(* Logix 5000 project; controller PLC_MCC1300_75F1 vendor 1 type 14 code 166 rev 32.11; software revision 32.04; part 81 of 83 *)
(* tags used below, declared in another part *)
   GP_OB_InitializeMain : GP_OB_Initialize;
   M302SpeedUp : MAC_SpeedUp;
   M307D_M1_DR : AXIS_CIP_DRIVE;
   M307E_M1_DR : AXIS_CIP_DRIVE;
   M307F_M1_DR : AXIS_CIP_DRIVE;
   M310_M1_DR_R1 : AXIS_CIP_DRIVE;
   M310_M2_DR_R2 : AXIS_CIP_DRIVE;
   M310_M3_DR_R3 : AXIS_CIP_DRIVE;
   TMP_dDirection : DINT;
   TMP_dTarget : DINT;
   TMP_rAcc : REAL;
   TMP_rDec : REAL;
   TMP_rSpeed : REAL;
   Z300_Conveyor : UDT_StandConv[29];
   Z300_Conveyor_IN_MOTION : MAC_Conveyor_ZC_IN_MOTION[29];
   Z300_Conveyor_OUT_MOTION : MAC_Conveyor_ZC_OUT_MOTION[29];
(* MotionLogic, continued *)

ROUTINE M307D_Motion   (* ladder *)
   // M307DM1
   0: NOP();
   1: XIC(Z300_Conveyor[18].OUTPUT_xDriveReset.0)MASR(M307D_M1_DR,Z300_Conveyor_OUT_MOTION[18].DR_MASR_M[0]);
   2: [XIC(Z300_Conveyor[18].OUTPUT_xDriveEnable.[0]) XIO(Z300_Conveyor_OUT_MOTION[18].DR_MSO_M[0].ER) MSO(M307D_M1_DR,Z300_Conveyor_OUT_MOTION[18].DR_MSO_M[0]) ,XIO(Z300_Conveyor_OUT_MOTION[18].DR_MSO_M[0].EN) OTU(Z300_Conveyor_OUT_MOTION[18].DR_MSO_M[0].ER) ,XIO(Z300_Conveyor[18].OUTPUT_xDriveEnable.[0]) OTU(Z300_Conveyor_OUT_MOTION[18].DR_MSO_M[0].EN) XIO(Z300_Conveyor_OUT_MOTION[18].DR_MSF_M[0].ER) MSF(M307D_M1_DR,Z300_Conveyor_OUT_MOTION[18].DR_MSF_M[0]) ,XIO(Z300_Conveyor_OUT_MOTION[18].DR_MSF_M[0].EN) OTU(Z300_Conveyor_OUT_MOTION[18].DR_MSF_M[0].ER) ];
   3: MUL(Z300_Conveyor[18].AUX_rgrAcc_m_s2[0],1000,TMP_rAcc)MUL(Z300_Conveyor[18].AUX_rgrDec_m_s2[0],1000,TMP_rDec)DIV(Z300_Conveyor[18].AUX_rgdRequestSpeed_mm_min[0],60,TMP_rSpeed);
   4: XIC(Z300_Conveyor[18].OS_xStartCount.0)OTU(Z300_Conveyor_IN_MOTION[18].DR_MAR_M[0].PC)OTU(Z300_Conveyor_IN_MOTION[18].DR_MRP_M[0].DN);
   5: [XIC(Z300_Conveyor[18].OUTPUT_xRun.0) MOV(0,TMP_dDirection) ,XIC(Z300_Conveyor[18].OUTPUT_xReverse.0) MOV(1,TMP_dDirection) ][XIO(Z300_Conveyor_IN_MOTION[18].DR_MAR_M[0].PC) ,XIO(Z300_Conveyor_IN_MOTION[18].DR_MRP_M[0].DN) ,XIO(Z300_Conveyor[18].OUTPUT_xPositioning.0) ]MAJ(M307D_M1_DR,Z300_Conveyor_OUT_MOTION[18].DR_MAJ_M[0],TMP_dDirection,TMP_rSpeed,Units per sec,TMP_rAcc,Units per sec2,TMP_rDec,Units per sec2,Trapezoidal,TMP_rAcc,TMP_rDec,Units per sec3,Enabled,Programmed,0,None);
   6: XIC(Z300_Conveyor[18].OS_xStartCount.0)MRP(M307D_M1_DR,Z300_Conveyor_OUT_MOTION[18].DR_MRP_M[0],Absolute,Actual,0);
   7: [XIC(Z300_Conveyor_IN_MOTION[18].DR_MRP_M[0].DN) XIC(Z300_Conveyor[18].OUTPUT_xPositioning.0) [XIC(Z300_Conveyor[18].tmON_PhFilter[0].DN) ,XIC(Z300_Conveyor_IN_MOTION[18].DR_MAR_M[0].EN) ] MAR(M307D_M1_DR,Z300_Conveyor_OUT_MOTION[18].DR_MAR_M[0],Negative_Edge,Disabled,0,0,1) ,XIO(Z300_Conveyor[18].OUTPUT_xPositioning.0) MDR(M307D_M1_DR,Z300_Conveyor_OUT_MOTION[18].DR_MDR_M[0],1) ];
   8: XIC(Z300_Conveyor[18].OUTPUT_xPositioning.0)XIC(Z300_Conveyor_IN_MOTION[18].DR_MAR_M[0].PC)DIV(Z300_Conveyor[18].AUX_rgdTarget_cmm[0],100,TMP_dTarget)ADD(TMP_dTarget,M307D_M1_DR.Registration1Position,TMP_dTarget)MAM(M307D_M1_DR,Z300_Conveyor_OUT_MOTION[18].DR_MAM_M[0],0,TMP_dTarget,TMP_rSpeed,Units per sec,TMP_rAcc,Units per sec2,TMP_rDec,Units per sec2,Trapezoidal,TMP_rAcc,TMP_rDec,Units per sec3,Enabled,Programmed,0,None,0,0);
   9: [XIC(Z300_Conveyor[18].OUTPUT_xChangeSpeed.0) ,XIC(M302SpeedUp.OS_xChangeAccDec) ,XIC(GP_OB_InitializeMain.OUT_xOs_200ms) ][XIO(Z300_Conveyor[18].OUTPUT_xReverse.0) ,XIC(Z300_Conveyor[18].OUTPUT_xReverse.0) MUL(TMP_rSpeed,-1.0,TMP_rSpeed) ]MCD(M307D_M1_DR,Z300_Conveyor_OUT_MOTION[18].DR_MCD_M[0],Jog,Yes,TMP_rSpeed,Yes,TMP_rAcc,Yes,TMP_rDec,No,TMP_rAcc,No,TMP_rDec,Units per sec,Units per sec2,Units per sec2,Units per sec3);
   10: XIO(Z300_Conveyor[18].OUTPUT_xRun.0)XIO(Z300_Conveyor[18].OUTPUT_xReverse.0)[XIC(Z300_Conveyor_IN_MOTION[18].DR_MAJ_M[0].IP) MAS(M307D_M1_DR,Z300_Conveyor_OUT_MOTION[18].DR_MASjog_M[0],Jog,Yes,TMP_rDec,Units per sec2,No,TMP_rDec,Units per sec3) ,XIC(Z300_Conveyor_IN_MOTION[18].DR_MAM_M[0].IP) MAS(M307D_M1_DR,Z300_Conveyor_OUT_MOTION[18].DR_MASpos_M[0],Move,Yes,TMP_rDec,Units per sec2,No,TMP_rDec,Units per sec3) ,XIO(Z300_Conveyor_IN_MOTION[18].DR_MAJ_M[0].IP) XIO(Z300_Conveyor_IN_MOTION[18].DR_MAM_M[0].IP) XIO(Z300_Conveyor_IN_MOTION[18].DR_MASjog_M[0].IP) XIO(Z300_Conveyor_IN_MOTION[18].DR_MASpos_M[0].IP) MAS(M307D_M1_DR,Z300_Conveyor_OUT_MOTION[18].DR_MASall_M[0],All,Yes,TMP_rDec,Units per sec2,No,TMP_rDec,Units per sec3) ];
END_ROUTINE

ROUTINE M307E_Motion   (* ladder *)
   // M307EM1
   0: NOP();
   1: XIC(Z300_Conveyor[19].OUTPUT_xDriveReset.0)MASR(M307E_M1_DR,Z300_Conveyor_OUT_MOTION[19].DR_MASR_M[0]);
   2: [XIC(Z300_Conveyor[19].OUTPUT_xDriveEnable.[0]) XIO(Z300_Conveyor_OUT_MOTION[19].DR_MSO_M[0].ER) MSO(M307E_M1_DR,Z300_Conveyor_OUT_MOTION[19].DR_MSO_M[0]) ,XIO(Z300_Conveyor_OUT_MOTION[19].DR_MSO_M[0].EN) OTU(Z300_Conveyor_OUT_MOTION[19].DR_MSO_M[0].ER) ,XIO(Z300_Conveyor[19].OUTPUT_xDriveEnable.[0]) OTU(Z300_Conveyor_OUT_MOTION[19].DR_MSO_M[0].EN) XIO(Z300_Conveyor_OUT_MOTION[19].DR_MSF_M[0].ER) MSF(M307E_M1_DR,Z300_Conveyor_OUT_MOTION[19].DR_MSF_M[0]) ,XIO(Z300_Conveyor_OUT_MOTION[19].DR_MSF_M[0].EN) OTU(Z300_Conveyor_OUT_MOTION[19].DR_MSF_M[0].ER) ];
   3: MUL(Z300_Conveyor[19].AUX_rgrAcc_m_s2[0],1000,TMP_rAcc)MUL(Z300_Conveyor[19].AUX_rgrDec_m_s2[0],1000,TMP_rDec)DIV(Z300_Conveyor[19].AUX_rgdRequestSpeed_mm_min[0],60,TMP_rSpeed);
   4: XIC(Z300_Conveyor[19].OS_xStartCount.0)OTU(Z300_Conveyor_IN_MOTION[19].DR_MAR_M[0].PC)OTU(Z300_Conveyor_IN_MOTION[19].DR_MRP_M[0].DN);
   5: [XIC(Z300_Conveyor[19].OUTPUT_xRun.0) MOV(0,TMP_dDirection) ,XIC(Z300_Conveyor[19].OUTPUT_xReverse.0) MOV(1,TMP_dDirection) ][XIO(Z300_Conveyor_IN_MOTION[19].DR_MAR_M[0].PC) ,XIO(Z300_Conveyor_IN_MOTION[19].DR_MRP_M[0].DN) ,XIO(Z300_Conveyor[19].OUTPUT_xPositioning.0) ]MAJ(M307E_M1_DR,Z300_Conveyor_OUT_MOTION[19].DR_MAJ_M[0],TMP_dDirection,TMP_rSpeed,Units per sec,TMP_rAcc,Units per sec2,TMP_rDec,Units per sec2,Trapezoidal,TMP_rAcc,TMP_rDec,Units per sec3,Enabled,Programmed,0,None);
   6: XIC(Z300_Conveyor[19].OS_xStartCount.0)MRP(M307E_M1_DR,Z300_Conveyor_OUT_MOTION[19].DR_MRP_M[0],Absolute,Actual,0);
   7: [XIC(Z300_Conveyor_IN_MOTION[19].DR_MRP_M[0].DN) XIC(Z300_Conveyor[19].OUTPUT_xPositioning.0) [XIC(Z300_Conveyor[19].tmON_PhFilter[0].DN) ,XIC(Z300_Conveyor_IN_MOTION[19].DR_MAR_M[0].EN) ] MAR(M307E_M1_DR,Z300_Conveyor_OUT_MOTION[19].DR_MAR_M[0],Negative_Edge,Disabled,0,0,1) ,XIO(Z300_Conveyor[19].OUTPUT_xPositioning.0) MDR(M307E_M1_DR,Z300_Conveyor_OUT_MOTION[19].DR_MDR_M[0],1) ];
   8: XIC(Z300_Conveyor[19].OUTPUT_xPositioning.0)XIC(Z300_Conveyor_IN_MOTION[19].DR_MAR_M[0].PC)DIV(Z300_Conveyor[19].AUX_rgdTarget_cmm[0],100,TMP_dTarget)ADD(TMP_dTarget,M307E_M1_DR.Registration1Position,TMP_dTarget)MAM(M307E_M1_DR,Z300_Conveyor_OUT_MOTION[19].DR_MAM_M[0],0,TMP_dTarget,TMP_rSpeed,Units per sec,TMP_rAcc,Units per sec2,TMP_rDec,Units per sec2,Trapezoidal,TMP_rAcc,TMP_rDec,Units per sec3,Enabled,Programmed,0,None,0,0);
   9: [XIC(Z300_Conveyor[19].OUTPUT_xChangeSpeed.0) ,XIC(M302SpeedUp.OS_xChangeAccDec) ,XIC(GP_OB_InitializeMain.OUT_xOs_200ms) ][XIO(Z300_Conveyor[19].OUTPUT_xReverse.0) ,XIC(Z300_Conveyor[19].OUTPUT_xReverse.0) MUL(TMP_rSpeed,-1.0,TMP_rSpeed) ]MCD(M307E_M1_DR,Z300_Conveyor_OUT_MOTION[19].DR_MCD_M[0],Jog,Yes,TMP_rSpeed,Yes,TMP_rAcc,Yes,TMP_rDec,No,TMP_rAcc,No,TMP_rDec,Units per sec,Units per sec2,Units per sec2,Units per sec3);
   10: XIO(Z300_Conveyor[19].OUTPUT_xRun.0)XIO(Z300_Conveyor[19].OUTPUT_xReverse.0)[XIC(Z300_Conveyor_IN_MOTION[19].DR_MAJ_M[0].IP) MAS(M307E_M1_DR,Z300_Conveyor_OUT_MOTION[19].DR_MASjog_M[0],Jog,Yes,TMP_rDec,Units per sec2,No,TMP_rDec,Units per sec3) ,XIC(Z300_Conveyor_IN_MOTION[19].DR_MAM_M[0].IP) MAS(M307E_M1_DR,Z300_Conveyor_OUT_MOTION[19].DR_MASpos_M[0],Move,Yes,TMP_rDec,Units per sec2,No,TMP_rDec,Units per sec3) ,XIO(Z300_Conveyor_IN_MOTION[19].DR_MAJ_M[0].IP) XIO(Z300_Conveyor_IN_MOTION[19].DR_MAM_M[0].IP) XIO(Z300_Conveyor_IN_MOTION[19].DR_MASjog_M[0].IP) XIO(Z300_Conveyor_IN_MOTION[19].DR_MASpos_M[0].IP) MAS(M307E_M1_DR,Z300_Conveyor_OUT_MOTION[19].DR_MASall_M[0],All,Yes,TMP_rDec,Units per sec2,No,TMP_rDec,Units per sec3) ];
END_ROUTINE

ROUTINE M307F_Motion   (* ladder *)
   // M307FM1
   0: NOP();
   1: XIC(Z300_Conveyor[20].OUTPUT_xDriveReset.0)MASR(M307F_M1_DR,Z300_Conveyor_OUT_MOTION[20].DR_MASR_M[0]);
   2: [XIC(Z300_Conveyor[20].OUTPUT_xDriveEnable.[0]) XIO(Z300_Conveyor_OUT_MOTION[20].DR_MSO_M[0].ER) MSO(M307F_M1_DR,Z300_Conveyor_OUT_MOTION[20].DR_MSO_M[0]) ,XIO(Z300_Conveyor_OUT_MOTION[20].DR_MSO_M[0].EN) OTU(Z300_Conveyor_OUT_MOTION[20].DR_MSO_M[0].ER) ,XIO(Z300_Conveyor[20].OUTPUT_xDriveEnable.[0]) OTU(Z300_Conveyor_OUT_MOTION[20].DR_MSO_M[0].EN) XIO(Z300_Conveyor_OUT_MOTION[20].DR_MSF_M[0].ER) MSF(M307F_M1_DR,Z300_Conveyor_OUT_MOTION[20].DR_MSF_M[0]) ,XIO(Z300_Conveyor_OUT_MOTION[20].DR_MSF_M[0].EN) OTU(Z300_Conveyor_OUT_MOTION[20].DR_MSF_M[0].ER) ];
   3: MUL(Z300_Conveyor[20].AUX_rgrAcc_m_s2[0],1000,TMP_rAcc)MUL(Z300_Conveyor[20].AUX_rgrDec_m_s2[0],1000,TMP_rDec)DIV(Z300_Conveyor[20].AUX_rgdRequestSpeed_mm_min[0],60,TMP_rSpeed);
   4: XIC(Z300_Conveyor[20].OS_xStartCount.0)OTU(Z300_Conveyor_IN_MOTION[20].DR_MAR_M[0].PC)OTU(Z300_Conveyor_IN_MOTION[20].DR_MRP_M[0].DN);
   5: [XIC(Z300_Conveyor[20].OUTPUT_xRun.0) MOV(0,TMP_dDirection) ,XIC(Z300_Conveyor[20].OUTPUT_xReverse.0) MOV(1,TMP_dDirection) ][XIO(Z300_Conveyor_IN_MOTION[20].DR_MAR_M[0].PC) ,XIO(Z300_Conveyor_IN_MOTION[20].DR_MRP_M[0].DN) ,XIO(Z300_Conveyor[20].OUTPUT_xPositioning.0) ]MAJ(M307F_M1_DR,Z300_Conveyor_OUT_MOTION[20].DR_MAJ_M[0],TMP_dDirection,TMP_rSpeed,Units per sec,TMP_rAcc,Units per sec2,TMP_rDec,Units per sec2,Trapezoidal,TMP_rAcc,TMP_rDec,Units per sec3,Enabled,Programmed,0,None);
   6: XIC(Z300_Conveyor[20].OS_xStartCount.0)MRP(M307F_M1_DR,Z300_Conveyor_OUT_MOTION[20].DR_MRP_M[0],Absolute,Actual,0);
   7: [XIC(Z300_Conveyor_IN_MOTION[20].DR_MRP_M[0].DN) XIC(Z300_Conveyor[20].OUTPUT_xPositioning.0) [XIC(Z300_Conveyor[20].tmON_PhFilter[0].DN) ,XIC(Z300_Conveyor_IN_MOTION[20].DR_MAR_M[0].EN) ] MAR(M307F_M1_DR,Z300_Conveyor_OUT_MOTION[20].DR_MAR_M[0],Negative_Edge,Disabled,0,0,1) ,XIO(Z300_Conveyor[20].OUTPUT_xPositioning.0) MDR(M307F_M1_DR,Z300_Conveyor_OUT_MOTION[20].DR_MDR_M[0],1) ];
   8: XIC(Z300_Conveyor[20].OUTPUT_xPositioning.0)XIC(Z300_Conveyor_IN_MOTION[20].DR_MAR_M[0].PC)DIV(Z300_Conveyor[20].AUX_rgdTarget_cmm[0],100,TMP_dTarget)ADD(TMP_dTarget,M307F_M1_DR.Registration1Position,TMP_dTarget)MAM(M307F_M1_DR,Z300_Conveyor_OUT_MOTION[20].DR_MAM_M[0],0,TMP_dTarget,TMP_rSpeed,Units per sec,TMP_rAcc,Units per sec2,TMP_rDec,Units per sec2,Trapezoidal,TMP_rAcc,TMP_rDec,Units per sec3,Enabled,Programmed,0,None,0,0);
   9: [XIC(Z300_Conveyor[20].OUTPUT_xChangeSpeed.0) ,XIC(M302SpeedUp.OS_xChangeAccDec) ,XIC(GP_OB_InitializeMain.OUT_xOs_200ms) ][XIO(Z300_Conveyor[20].OUTPUT_xReverse.0) ,XIC(Z300_Conveyor[20].OUTPUT_xReverse.0) MUL(TMP_rSpeed,-1.0,TMP_rSpeed) ]MCD(M307F_M1_DR,Z300_Conveyor_OUT_MOTION[20].DR_MCD_M[0],Jog,Yes,TMP_rSpeed,Yes,TMP_rAcc,Yes,TMP_rDec,No,TMP_rAcc,No,TMP_rDec,Units per sec,Units per sec2,Units per sec2,Units per sec3);
   10: XIO(Z300_Conveyor[20].OUTPUT_xRun.0)XIO(Z300_Conveyor[20].OUTPUT_xReverse.0)[XIC(Z300_Conveyor_IN_MOTION[20].DR_MAJ_M[0].IP) MAS(M307F_M1_DR,Z300_Conveyor_OUT_MOTION[20].DR_MASjog_M[0],Jog,Yes,TMP_rDec,Units per sec2,No,TMP_rDec,Units per sec3) ,XIC(Z300_Conveyor_IN_MOTION[20].DR_MAM_M[0].IP) MAS(M307F_M1_DR,Z300_Conveyor_OUT_MOTION[20].DR_MASpos_M[0],Move,Yes,TMP_rDec,Units per sec2,No,TMP_rDec,Units per sec3) ,XIO(Z300_Conveyor_IN_MOTION[20].DR_MAJ_M[0].IP) XIO(Z300_Conveyor_IN_MOTION[20].DR_MAM_M[0].IP) XIO(Z300_Conveyor_IN_MOTION[20].DR_MASjog_M[0].IP) XIO(Z300_Conveyor_IN_MOTION[20].DR_MASpos_M[0].IP) MAS(M307F_M1_DR,Z300_Conveyor_OUT_MOTION[20].DR_MASall_M[0],All,Yes,TMP_rDec,Units per sec2,No,TMP_rDec,Units per sec3) ];
END_ROUTINE

ROUTINE M310_Motion   (* ladder *)
   // M310M1
   0: NOP();
   1: XIC(Z300_Conveyor[22].OUTPUT_xDriveReset.0)MASR(M310_M1_DR_R1,Z300_Conveyor_OUT_MOTION[22].DR_MASR_M[0]);
   2: [XIC(Z300_Conveyor[22].OUTPUT_xDriveEnable.[0]) XIO(Z300_Conveyor_OUT_MOTION[22].DR_MSO_M[0].ER) MSO(M310_M1_DR_R1,Z300_Conveyor_OUT_MOTION[22].DR_MSO_M[0]) ,XIO(Z300_Conveyor_OUT_MOTION[22].DR_MSO_M[0].EN) OTU(Z300_Conveyor_OUT_MOTION[22].DR_MSO_M[0].ER) ,XIO(Z300_Conveyor[22].OUTPUT_xDriveEnable.[0]) OTU(Z300_Conveyor_OUT_MOTION[22].DR_MSO_M[0].EN) XIO(Z300_Conveyor_OUT_MOTION[22].DR_MSF_M[0].ER) MSF(M310_M1_DR_R1,Z300_Conveyor_OUT_MOTION[22].DR_MSF_M[0]) ,XIO(Z300_Conveyor_OUT_MOTION[22].DR_MSF_M[0].EN) OTU(Z300_Conveyor_OUT_MOTION[22].DR_MSF_M[0].ER) ];
   3: MUL(Z300_Conveyor[22].AUX_rgrAcc_m_s2[0],1000,TMP_rAcc)MUL(Z300_Conveyor[22].AUX_rgrDec_m_s2[0],1000,TMP_rDec)DIV(Z300_Conveyor[22].AUX_rgdRequestSpeed_mm_min[0],60,TMP_rSpeed);
   4: XIC(Z300_Conveyor[22].OS_xStartCount.0)OTU(Z300_Conveyor_IN_MOTION[22].DR_MAR_M[0].PC)OTU(Z300_Conveyor_IN_MOTION[22].DR_MRP_M[0].DN);
   5: [XIC(Z300_Conveyor[22].OUTPUT_xRun.0) MOV(0,TMP_dDirection) ,XIC(Z300_Conveyor[22].OUTPUT_xReverse.0) MOV(1,TMP_dDirection) ][XIO(Z300_Conveyor_IN_MOTION[22].DR_MAR_M[0].PC) ,XIO(Z300_Conveyor_IN_MOTION[22].DR_MRP_M[0].DN) ,XIO(Z300_Conveyor[22].OUTPUT_xPositioning.0) ]MAJ(M310_M1_DR_R1,Z300_Conveyor_OUT_MOTION[22].DR_MAJ_M[0],TMP_dDirection,TMP_rSpeed,Units per sec,TMP_rAcc,Units per sec2,TMP_rDec,Units per sec2,Trapezoidal,TMP_rAcc,TMP_rDec,Units per sec3,Enabled,Programmed,0,None);
   6: XIC(Z300_Conveyor[22].OS_xStartCount.0)MRP(M310_M1_DR_R1,Z300_Conveyor_OUT_MOTION[22].DR_MRP_M[0],Absolute,Actual,0);
   7: [XIC(Z300_Conveyor_IN_MOTION[22].DR_MRP_M[0].DN) XIC(Z300_Conveyor[22].OUTPUT_xPositioning.0) [XIC(Z300_Conveyor[22].tmON_PhFilter[0].DN) ,XIC(Z300_Conveyor_IN_MOTION[22].DR_MAR_M[0].EN) ] MAR(M310_M1_DR_R1,Z300_Conveyor_OUT_MOTION[22].DR_MAR_M[0],Negative_Edge,Disabled,0,0,1) ,XIO(Z300_Conveyor[22].OUTPUT_xPositioning.0) MDR(M310_M1_DR_R1,Z300_Conveyor_OUT_MOTION[22].DR_MDR_M[0],1) ];
   8: XIC(Z300_Conveyor[22].OUTPUT_xPositioning.0)XIC(Z300_Conveyor_IN_MOTION[22].DR_MAR_M[0].PC)DIV(Z300_Conveyor[22].AUX_rgdTarget_cmm[0],100,TMP_dTarget)ADD(TMP_dTarget,M310_M1_DR_R1.Registration1Position,TMP_dTarget)MAM(M310_M1_DR_R1,Z300_Conveyor_OUT_MOTION[22].DR_MAM_M[0],0,TMP_dTarget,TMP_rSpeed,Units per sec,TMP_rAcc,Units per sec2,TMP_rDec,Units per sec2,Trapezoidal,TMP_rAcc,TMP_rDec,Units per sec3,Enabled,Programmed,0,None,0,0);
   9: [XIC(Z300_Conveyor[22].OUTPUT_xChangeSpeed.0) ,XIC(M302SpeedUp.OS_xChangeAccDec) ,XIC(GP_OB_InitializeMain.OUT_xOs_200ms) ][XIO(Z300_Conveyor[22].OUTPUT_xReverse.0) ,XIC(Z300_Conveyor[22].OUTPUT_xReverse.0) MUL(TMP_rSpeed,-1.0,TMP_rSpeed) ]MCD(M310_M1_DR_R1,Z300_Conveyor_OUT_MOTION[22].DR_MCD_M[0],Jog,Yes,TMP_rSpeed,Yes,TMP_rAcc,Yes,TMP_rDec,No,TMP_rAcc,No,TMP_rDec,Units per sec,Units per sec2,Units per sec2,Units per sec3);
   10: XIO(Z300_Conveyor[22].OUTPUT_xRun.0)XIO(Z300_Conveyor[22].OUTPUT_xReverse.0)[XIC(Z300_Conveyor_IN_MOTION[22].DR_MAJ_M[0].IP) MAS(M310_M1_DR_R1,Z300_Conveyor_OUT_MOTION[22].DR_MASjog_M[0],Jog,Yes,TMP_rDec,Units per sec2,No,TMP_rDec,Units per sec3) ,XIC(Z300_Conveyor_IN_MOTION[22].DR_MAM_M[0].IP) MAS(M310_M1_DR_R1,Z300_Conveyor_OUT_MOTION[22].DR_MASpos_M[0],Move,Yes,TMP_rDec,Units per sec2,No,TMP_rDec,Units per sec3) ,XIO(Z300_Conveyor_IN_MOTION[22].DR_MAJ_M[0].IP) XIO(Z300_Conveyor_IN_MOTION[22].DR_MAM_M[0].IP) XIO(Z300_Conveyor_IN_MOTION[22].DR_MASjog_M[0].IP) XIO(Z300_Conveyor_IN_MOTION[22].DR_MASpos_M[0].IP) MAS(M310_M1_DR_R1,Z300_Conveyor_OUT_MOTION[22].DR_MASall_M[0],All,Yes,TMP_rDec,Units per sec2,No,TMP_rDec,Units per sec3) ];
   // M310M2
   11: NOP();
   12: XIC(Z300_Conveyor[23].OUTPUT_xDriveReset.0)MASR(M310_M2_DR_R2,Z300_Conveyor_OUT_MOTION[23].DR_MASR_M[0]);
   13: [XIC(Z300_Conveyor[23].OUTPUT_xDriveEnable.[0]) XIO(Z300_Conveyor_OUT_MOTION[23].DR_MSO_M[0].ER) MSO(M310_M2_DR_R2,Z300_Conveyor_OUT_MOTION[23].DR_MSO_M[0]) ,XIO(Z300_Conveyor_OUT_MOTION[23].DR_MSO_M[0].EN) OTU(Z300_Conveyor_OUT_MOTION[23].DR_MSO_M[0].ER) ,XIO(Z300_Conveyor[23].OUTPUT_xDriveEnable.[0]) OTU(Z300_Conveyor_OUT_MOTION[23].DR_MSO_M[0].EN) XIO(Z300_Conveyor_OUT_MOTION[23].DR_MSF_M[0].ER) MSF(M310_M2_DR_R2,Z300_Conveyor_OUT_MOTION[23].DR_MSF_M[0]) ,XIO(Z300_Conveyor_OUT_MOTION[23].DR_MSF_M[0].EN) OTU(Z300_Conveyor_OUT_MOTION[23].DR_MSF_M[0].ER) ];
   14: MUL(Z300_Conveyor[23].AUX_rgrAcc_m_s2[0],1000,TMP_rAcc)MUL(Z300_Conveyor[23].AUX_rgrDec_m_s2[0],1000,TMP_rDec)DIV(Z300_Conveyor[23].AUX_rgdRequestSpeed_mm_min[0],60,TMP_rSpeed);
   15: XIC(Z300_Conveyor[23].OS_xStartCount.0)OTU(Z300_Conveyor_IN_MOTION[23].DR_MAR_M[0].PC)OTU(Z300_Conveyor_IN_MOTION[23].DR_MRP_M[0].DN);
   16: [XIC(Z300_Conveyor[23].OUTPUT_xRun.0) MOV(0,TMP_dDirection) ,XIC(Z300_Conveyor[23].OUTPUT_xReverse.0) MOV(1,TMP_dDirection) ][XIO(Z300_Conveyor_IN_MOTION[23].DR_MAR_M[0].PC) ,XIO(Z300_Conveyor_IN_MOTION[23].DR_MRP_M[0].DN) ,XIO(Z300_Conveyor[23].OUTPUT_xPositioning.0) ]MAJ(M310_M2_DR_R2,Z300_Conveyor_OUT_MOTION[23].DR_MAJ_M[0],TMP_dDirection,TMP_rSpeed,Units per sec,TMP_rAcc,Units per sec2,TMP_rDec,Units per sec2,Trapezoidal,TMP_rAcc,TMP_rDec,Units per sec3,Enabled,Programmed,0,None);
   17: XIC(Z300_Conveyor[23].OS_xStartCount.0)MRP(M310_M2_DR_R2,Z300_Conveyor_OUT_MOTION[23].DR_MRP_M[0],Absolute,Actual,0);
   18: [XIC(Z300_Conveyor_IN_MOTION[23].DR_MRP_M[0].DN) XIC(Z300_Conveyor[23].OUTPUT_xPositioning.0) [XIC(Z300_Conveyor[23].tmON_PhFilter[0].DN) ,XIC(Z300_Conveyor_IN_MOTION[23].DR_MAR_M[0].EN) ] MAR(M310_M2_DR_R2,Z300_Conveyor_OUT_MOTION[23].DR_MAR_M[0],Negative_Edge,Disabled,0,0,1) ,XIO(Z300_Conveyor[23].OUTPUT_xPositioning.0) MDR(M310_M2_DR_R2,Z300_Conveyor_OUT_MOTION[23].DR_MDR_M[0],1) ];
   19: XIC(Z300_Conveyor[23].OUTPUT_xPositioning.0)XIC(Z300_Conveyor_IN_MOTION[23].DR_MAR_M[0].PC)DIV(Z300_Conveyor[23].AUX_rgdTarget_cmm[0],100,TMP_dTarget)ADD(TMP_dTarget,M310_M2_DR_R2.Registration1Position,TMP_dTarget)MAM(M310_M2_DR_R2,Z300_Conveyor_OUT_MOTION[23].DR_MAM_M[0],0,TMP_dTarget,TMP_rSpeed,Units per sec,TMP_rAcc,Units per sec2,TMP_rDec,Units per sec2,Trapezoidal,TMP_rAcc,TMP_rDec,Units per sec3,Enabled,Programmed,0,None,0,0);
   20: [XIC(Z300_Conveyor[23].OUTPUT_xChangeSpeed.0) ,XIC(M302SpeedUp.OS_xChangeAccDec) ,XIC(GP_OB_InitializeMain.OUT_xOs_200ms) ][XIO(Z300_Conveyor[23].OUTPUT_xReverse.0) ,XIC(Z300_Conveyor[23].OUTPUT_xReverse.0) MUL(TMP_rSpeed,-1.0,TMP_rSpeed) ]MCD(M310_M2_DR_R2,Z300_Conveyor_OUT_MOTION[23].DR_MCD_M[0],Jog,Yes,TMP_rSpeed,Yes,TMP_rAcc,Yes,TMP_rDec,No,TMP_rAcc,No,TMP_rDec,Units per sec,Units per sec2,Units per sec2,Units per sec3);
   21: XIO(Z300_Conveyor[23].OUTPUT_xRun.0)XIO(Z300_Conveyor[23].OUTPUT_xReverse.0)[XIC(Z300_Conveyor_IN_MOTION[23].DR_MAJ_M[0].IP) MAS(M310_M2_DR_R2,Z300_Conveyor_OUT_MOTION[23].DR_MASjog_M[0],Jog,Yes,TMP_rDec,Units per sec2,No,TMP_rDec,Units per sec3) ,XIC(Z300_Conveyor_IN_MOTION[23].DR_MAM_M[0].IP) MAS(M310_M2_DR_R2,Z300_Conveyor_OUT_MOTION[23].DR_MASpos_M[0],Move,Yes,TMP_rDec,Units per sec2,No,TMP_rDec,Units per sec3) ,XIO(Z300_Conveyor_IN_MOTION[23].DR_MAJ_M[0].IP) XIO(Z300_Conveyor_IN_MOTION[23].DR_MAM_M[0].IP) XIO(Z300_Conveyor_IN_MOTION[23].DR_MASjog_M[0].IP) XIO(Z300_Conveyor_IN_MOTION[23].DR_MASpos_M[0].IP) MAS(M310_M2_DR_R2,Z300_Conveyor_OUT_MOTION[23].DR_MASall_M[0],All,Yes,TMP_rDec,Units per sec2,No,TMP_rDec,Units per sec3) ];
   // M310M2
   22: NOP();
   23: XIC(Z300_Conveyor[24].OUTPUT_xDriveReset.0)MASR(M310_M3_DR_R3,Z300_Conveyor_OUT_MOTION[24].DR_MASR_M[0]);
